FUNCTION_BLOCK "LKinCtrl_MC_ExecuteKinMotionCmd"   // FB35003, SCL
TITLE = LKinCtrl_ExecuteKinMotinCmd
{ S7_Optimized_Access := 'TRUE' }
AUTHOR : tech.team.motioncontrol@siemens.com
FAMILY : LKinCtrl
VERSION : 3.0
// FB executing single motion commands for TO_Kinematics. 
// - handling internal motion command instances
// - managing MotionQueue to be full, but not overloaded
// - providing status information on execution status
   VAR_INPUT
      execute : Bool;   // rising edge starts action once
      interrupt : Bool;   // trigger GroupInterrupt [interrupt input of FB_MovePath]
      continueMotion : Bool;   // trigger GroupContinue [no use in FB_MovePath] (used for FB_ExecutePathMotion stand alone)
      stop : Bool;   // trigger GroupStop [stop input of FB_MovePath]
      stopMode : DInt;   // MC_GroupStop dynamics; 0: stop with dynamics of active motion job; 1: stop with maximum kinematics dynamics (dynamics adaption still effective)
      reset : Bool;   // reset FB / acknowledge errors [reset input of FB_MovePath]
      writtenActiveCmdNo : DInt;   // last active cmdNo handled by FB MovePath
      conveyorConfiguration : Array[1.."LKINCTRL_NO_OF_CONVEYOR"] of "LKinCtrl_typeConveyorConfiguration";   // conveyor configuration / Conveyor configuration
   END_VAR
   VAR_OUTPUT
      done : Bool;   // TRUE: Commanded functionality has been completed successfully
      busy : Bool;   // TRUE: FB is not finished and new output values can be expected
      active : Bool;   // FB in control of axesGroup / kinematic in motion
      error : Bool;   // TRUE: An error occurred during the execution of the FB
      commandAborted : Bool;   // TRUE: Commanded functionality has been aborted by another command
      activePathDataName : String["LKINCTRL_LENGTH_OF_PATHDATA_NAME"];   // name of actual PathData
      activePathDataIdentifier : USInt;   // identifier number of actual PathData
      activeCmdNo : DInt;   // number of actual PathData set number
      cmdExecuted : Bool;   // actual pathData cmd executed to MotionQueue
      remainingDistanceActCmd : LReal;   // remainingDistance of active motionCommand
      waitTimeActive : Bool;   // TRUE: waitTime active in FB
      diagnostics : "LKinCtrl_typeExecuteKinMotionCmdDiagnostics";   // Diagnostics information of FB
   END_VAR
   VAR_IN_OUT
      pathDataElementPreBuf : "LKinCtrl_typePathDataElement_PreBuf";   // reference to the PathData element to be executed by FB_ExecuteKinMotionCmd
      to_Kinematics : TO_Kinematics;   // reference to the axesGroup
   END_VAR
   VAR
      statExecuteOld : Bool;   // old value of 'execute' input for edge detection
      statStopOld : Bool;   // old value of 'stop' input for edge detection
      statInterruptOld : Bool;   // old value of 'interrupt' input for edge detection
      statContinueMotionOld : Bool;   // old value of 'continueMotion' input for edge detection
      statResetOld : Bool;   // old value of 'reset' input for edge detection
      statDone : Bool;   // static value for output 'done'
      statBusy : Bool;   // static value for output 'busy'
      statCommandAborted : Bool;   // static value for output 'commandAborted'
      statActive : Bool;   // static value for output 'active'
      statActiveCmdNo : DInt;   // static value for output 'activeCmdNo'
      statWaitTimeActive : Bool;   // static value for output 'waitTimeActive'
      statWaitTime : Time;   // static time storage for time to wait for during wait time
      statError : Bool;   // static value for output 'error'
      statStatus : Word := 16#7000;   // static value for output 'status'
      statSubfunctionStatus : Word;   // Status or return value of called FBs, FCs and system blocks
      statFBState : Int := 0;   // State in the state machine of the FB
      statStateMachine : Int;   // static state machine status
      statDebugState : Bool;   // debug state machine by single steps
      statDebugFaultyValue : Int;   // debugging static for development only
      statDebugMessage : String;   // debugging string for development only
      statCmdExecuted : Bool;   // static value for output 'cmdExecuted'
      statExecWaitTime : Bool;   // execute flag for triggering wait time
      statExecFlagOnly : Bool;   // 'execute' flag for flagOnly dummy command
      statExecGroupInterrupt : Bool;   // execute flag for triggering MC_GroupInterrupt
      statExecGroupContinue : Bool;   // execute flag for triggering MC_GroupContinue
      statExecGroupStop : Bool;   // execute flag for triggering MC_GroupStop
      statExternalStopDetected : Bool;   // static storing informatioin on external stop being triggered
      statExecuteFlagOnlyCmd : Bool;   // static 'trigger' for execution of flag only cmd
      statStartCmdIsFlagOnly : Bool;   // static to store information that first command in PathData is flag only command
      statCmdIsMotionCmd : Bool;   // static containing cmd category; TRUE: motion cmd; FALSE: non-motion cmd
      statFBCounterLin : Int := 1;   // counter for organization of used linear motion FB instances
      statFBCounterCirc : Int := 1;   // counter for organization of used circular motion FB instances
      statFBCounterMoveDir : Int := 1;   // counter for organization of used move direct motion FB instances
      statFBCounterTrackConv : Int := 1;   // counter for organization of used conveyor tracking FB instances / counter for organization of used move direct motion FB instances
      statCoordSystemOld : DInt := 0;   // static storing old coordSystem information
      statLinkConstellation : DInt;   // static storing the link constellation
      statActualTrackedOCS : SInt;   // actually tracked OCS from kinematics
      statOCSInSync : SInt;   // OCS which is or will be syncrhonized to
      statBlendingRadius : LReal;   // calculated blending radius for SPTP commands
      statOCSInTracking : Array[1..3] of Bool;   // signalizes if a OCS is or will be used for tracking
      statLastPos : Array[1..4] of LReal;   // static for last TO_Kinematic position (for conversion relative to absolute motion)
      statAbsolutePosition : Array[1..4] of LReal;   // flag for AbsoultePosition of linear command to be changed internally (for conversion relative to absolute motion)
      statAuxPoint : Array[1..3] of LReal;   // flag for AuxPoint of circular command to be changed internally (for conversion relative to absolute motion)
      statEndPoint : Array[1..4] of LReal;   // flag for last EndPoint of circular command to be changed internally (for conversion relative to absolute motion)
      statExecLinCmds : Array[1..#LKINCTRL_MAX_NUMBER_OF_CMDS_LIN] of Bool;   // array of execute flags for triggering linear motion command FBs
      statExecCircCmds : Array[1..#LKINCTRL_MAX_NUMBER_OF_CMDS_CIRC] of Bool;   // array of execute flags for triggering circular motion command FBs
      statExecMoveDirectCmds : Array[1..#LKINCTRL_MAX_NUMBER_OF_CMDS_MOVEDIRECT] of Bool;   // array of execute flags for triggering move direct motion command FBs
      statExecTrackConv : Array[1..#LKINCTRL_MAX_NUMBER_OF_CMDS_TRACKCONV] of Bool;   // array of execute flags for triggering conveyor tracking command FBs / array of execute flags for triggering linear motion command FBs
      statConveyorBeltAxis : Array[1..#LKINCTRL_MAX_NUMBER_OF_CMDS_TRACKCONV] of DB_ANY;   // array of conveyor belt axes to be used at the instances
      statOCSFrames : Array[1..3] of "LKinCtrl_typeFrame";   // array of OCS frames
      statEmptyDiagnostics : "LKinCtrl_typeExecuteKinMotionCmdDiagnostics";   // empty diagnostics information (for initialization purposes only)
      statStoreExecuteBuffer : Struct   // struct for assignment of motion command FB instances PathData set specific data (setNo, PathDataNo)
         writeBufferElement : Int := 1;   // flag for set to be executed to MotionQueue in ExecuteBuffer struct
         activeBufferElement : Int := 1;   // flag for active set in ExecuteBuffer struct
         lastBufferElement : Int := 20;
         bufferElement : Array[1..#LKINCTRL_EXECUTEBUFFER_LENGTH] of Struct   // assignment of motion command FB instances PathData set specific data (setNo, PathDataNo)
            pathDataName : String["LKINCTRL_LENGTH_OF_PATHDATA_NAME"];
            pathDataIdentifier : USInt;
            setNumber : DInt;
            MotionFBNo : Int;
         END_STRUCT;
      END_STRUCT;
      statDebugExecCmdLogger : Struct   // command logger structure to store all executed commands (to MotionQueue), never deleted
         loggerElement : Array[1..#CONST_LENGTH_DATALOGGER] of Struct   // logger array storing executed commands and specific debug data
            executedCmd : "LKinCtrl_typeCmdLoggerElement";   // command
            executeBufferElement : Int;   // statStoreExecuteBuffer element number
            assignedMotionFB : Int;   // MC instance assigned
            timeStamp : Date_And_Time;   // time stamp of execution time of logged command
         END_STRUCT;
         writeCmdLoggerElement : Int := 1;   // pointer for writing logger element; incremented after writing ==> value -1 is last written element
         activeCmdLoggerElement : Int := 1;   // pointing on active cmd in command logger; showing active element during execution ==> after SUCCESSFUL completion of path incrementation ==> value -1 is last active element
      END_STRUCT;
      instMC_MoveLinAbs : Array[1..#LKINCTRL_MAX_NUMBER_OF_CMDS_LIN] of MC_MOVELINEARABSOLUTE;   // multi instance array MC_MoveLinearAbsoulte
      instMC_MoveCircAbs : Array[1..#LKINCTRL_MAX_NUMBER_OF_CMDS_CIRC] of MC_MOVECIRCULARABSOLUTE;   // multi instance array MC_MoveCircularAbsoulte
      instMC_MoveDirectAbs : Array[1..#LKINCTRL_MAX_NUMBER_OF_CMDS_MOVEDIRECT] of MC_MOVEDIRECTABSOLUTE;   // multi instance array MC_MoveDirectAbsoulte
      instMC_GROUPINTERRUPT : MC_GROUPINTERRUPT;   // multi instance MC_GroupInterrupt
      instMC_GROUPSTOP : MC_GROUPSTOP;   // multi instance FB MC_GroupStop
      instMC_GROUPCONTINUE : MC_GROUPCONTINUE;   // multi instance FB MC_GroupContinue
      instMC_KinematicsTransformation : MC_KINEMATICSTRANSFORMATION;   // multi instance FB MC_KinematicsTransformation
      instMC_InverseKinematicsTransformation : MC_INVERSEKINEMATICSTRANSFORMATION;   // multi instance FB MC_InverseKinematicsTransformation
      instMC_TrackConveyor : Array[1..3] of MC_TRACKCONVEYORBELT;   // multi instance FB MC_TrackConveyorBelt
      instIEC_Timer_waitTime : TON_TIME;   // multi instance TIMER_ON for wait times
   END_VAR
   VAR_TEMP
      tempExecute : Bool;   // Temporary value for input 'execute'
      tempStop : Bool;   // Temporary value for input 'stop'
      tempStopMode : DInt;   // Temporary value for input 'stopMode'
      tempInterrupt : Bool;   // Temporary value for input 'interrupt'
      tempContinueMotion : Bool;   // Temporary value for input 'continueMotion'
      tempReset : Bool;   // Temporary value for input 'reset'
      tempPosElemCtr : Int;   // Temporary counter variable
      tempCtr : Int;   // Temporary counter variable
      tempFBInstCtr : Int;   // Temporary counter variable
      tempMCActive : Bool;   // Temporary value to signal active MC instance
      tempMCBusy : Bool;   // Temporary value to signal busy MC instance
      tempRetVal : Int;   // Temporary return value
      tempRetValWord : Word;   // Temporary return value
      tempCmdType : Int;   // Temporary variable for type of command
      tempActiveInstance : Int;   // Temporary variable for active MC instance
      tempCmdDone : Bool;   // Temporary bit to signal done of MC instance
      tempCalc : Array[1..4] of LReal;   // Temporary calculation variable
      tempBlending : Array[1..4] of LReal;   // Temporary calculation variable
   END_VAR
   VAR CONSTANT
      NO_PROCESSING : Int := 0;   // FB_ExecutePathMotion state machine constant
      RESETTING : Int := 5;   // FB_ExecutePathMotion state machine constant
      RECEIVE_CMD : Int := 10;   // FB_ExecutePathMotion state machine constant
      CMD_CALC_SELECT : Int := 30;   // FB_ExecutePathMotion state machine constant
      EXEC_LIN : Int := 40;   // FB_ExecutePathMotion state machine constant
      EXEC_CIRC : Int := 41;   // FB_ExecutePathMotion state machine constant
      EXEC_MOVE_DIRECT : Int := 42;   // FB_ExecutePathMotion state machine constant
      EXEC_TRACK_CONV : Int := 43;   // FB_ExecutePathMotion state machine constant
      EXEC_SET_WS_ZONE : Int := 49;   // FB_ExecutePathMotion state machine constant
      EXEC_FLAG_ONLY : Int := 55;   // FB_ExecutePathMotion state machine constant
      EXEC_WAIT_TIME : Int := 57;   // FB_ExecutePathMotion state machine constant
      WAITING_TIME : Int := 58;   // FB_ExecutePathMotion state machine constant
      QUEUE_BUSY : Int := 60;   // FB_ExecutePathMotion state machine constant
      INTERRUPTING : Int := 70;   // FB_ExecutePathMotion state machine constant
      INTERRUPTED : Int := 75;   // FB_ExecutePathMotion state machine constant
      CONTINUEING : Int := 77;   // FB_ExecutePathMotion state machine constant
      CONTINUED : Int := 78;   // FB_ExecutePathMotion state machine constant
      STOPPING : Int := 80;   // FB_ExecutePathMotion state machine constant
      STOPPED_STATE : Int := 85;   // FB_ExecutePathMotion state machine constant
      DESYNC_CONVEYOR : Int := 86;   // FB_ExecutePathMotion state machine constant
      ERROR_STATE : Int := 90;   // FB_ExecutePathMotion state machine constant
      LKINCTRL_MAX_NUMBER_OF_CMDS_LIN : Int := 12;   // max number of MC_MoveLinearAbsolute FB instances
      LKINCTRL_MAX_NUMBER_OF_CMDS_CIRC : Int := 12;   // max number of MC_MoveCircularAbsolute FB instances
      LKINCTRL_MAX_NUMBER_OF_CMDS_MOVEDIRECT : Int := 12;   // max number of MC_MoveDirectAbsolute FB instances
      LKINCTRL_MAX_NUMBER_OF_CMDS_TRACKCONV : Int := 3;   // max number of MC_TrackConveyorBelt FB instances
      LKINCTRL_EXECUTEBUFFER_LENGTH : Int := 12;   // length of internal buffer (needs to be set to same value as LKINCTRL_MAX_NUMBER_OF_CMDS_LIN)
      STATUS_NO_ERROR : Word := 16#0000;   // status no error
      STATUS_NO_CALL : Word := 16#7000;   // No job being currently processed
      STATUS_FIRST_CALL : Word := 16#7001;   // First call after incoming new job (rising edge 'execute')
      STATUS_SUBSEQUENT_CALL : Word := 16#7002;   // Subsequent call during active processing without further details
      STATUS_CMD_EXECUTED : Word := 16#7010;   // status command executed to MotionQueue
      STATUS_PATHMOTION_RUNNING : Word := 16#7100;   // status path motion running
      STATUS_PATHMOTION_INTERRUPTING : Word := 16#7101;   // status path motion interrupting
      STATUS_PATHMOTION_INTERRUPTED : Word := 16#7102;   // status path motion interrupted
      STATUS_PATHMOTION_STOPPING : Word := 16#7103;   // status path motion stopping
      STATUS_COMMAND_ABORTED : Word := 16#7104;   // commanded functionality has been aborted by another command
      STATUS_PATHMOTION_CONTINUEING : Word := 16#7105;   // status path motion continueing
      STATUS_FB_RESETTING : Word := 16#7106;   // status FB reset
      STATUS_WAIT_TIME_ACTIVE : Word := 16#7107;   // status wait time active
      STATUS_WAIT_TIME_FINISHED : Word := 16#7108;   // status wait time finished
      STATUS_PATHMOTION_EXT_STOPPING : Word := 16#7109;   // status external stop active
      STATUS_PATHMOTION_BUFFER_BUSY : Word := 16#7111;   // status motionQueue full / buffer busy
      STATUS_PATHMOTION_FINISHED : Word := 16#7110;   // status path motion finished / end of path position reached
      STATUS_DESYNC_CONVEYOR : Word := 16#7112;   // status desync from conveyor with motion command
      ERR_UNDEFINED_STATE : Word := 16#8600;   // error due to an undefined state in state machine
      ERR_GROUPINTERRUPT_FAILED : Word := 16#8242;   // error MC_GroupInterrupt failed
      ERR_GROUPCONTINUE_FAILED : Word := 16#8243;   // error MC_GroupContinue failed
      ERR_GROUPSTOP_FAILED : Word := 16#8244;   // error MC_GroupStop failed
      ERR_TO_KINEMATIC_ERROR : Word := 16#8245;   // error in TO_Kinematic
      ERR_LINEAR_CMD : Word := 16#8246;   // error MC_MoveLinear failed
      ERR_CIRCULAR_CMD : Word := 16#8247;   // error MC_MoveCircular failed
      ERR_CMD_PARAMETER : Word := 16#8248;   // error command parametrization
      ERR_CALC_CIRC_CMD : Word := 16#8249;   // error circular command conversion: arc calculation
      ERR_MOVEDIRECT_CMD : Word := 16#8250;   // error MC_MoveDirect failed
      ERR_TRACKCONVEYOR_CMD : Word := 16#8251;   // error MC_TrackConveyorBelt failed
      ERR_DESYNC_RELATIVE : Word := 16#8252;   // error due to relative command used for desync conveyor
      ERR_CONVEYOR_CONFIGURATION : Word := 16#8253;   // error due to invalid conveyor configuration
      CONST_LENGTH_DATALOGGER : Int := 15;   // length of internal data logger
      SPTP_REMAINING_DIST : Bool := FALSE;   // TRUE: Caclulate own RemainingDistance for SPTP / FALSE: Use ExecutionTimeStatus
      SPTP_APPROX_BLENDING : Bool := FALSE;   // TRUE: When remDistance is calculated also approximate blending distance / FALSE: Set blending is not regarded on calculation
   END_VAR
   // statStoreExecuteBuffer.bufferElement[12].MotionFBNo := -1;
   // statStoreExecuteBuffer.bufferElement[11].MotionFBNo := -1;
   // statStoreExecuteBuffer.bufferElement[10].MotionFBNo := -1;
   // statStoreExecuteBuffer.bufferElement[9].MotionFBNo := -1;
   // statStoreExecuteBuffer.bufferElement[8].MotionFBNo := -1;
   // statStoreExecuteBuffer.bufferElement[7].MotionFBNo := -1;
   // statStoreExecuteBuffer.bufferElement[6].MotionFBNo := -1;
   // statStoreExecuteBuffer.bufferElement[5].MotionFBNo := -1;
   // statStoreExecuteBuffer.bufferElement[4].MotionFBNo := -1;
   // statStoreExecuteBuffer.bufferElement[3].MotionFBNo := -1;
   // statStoreExecuteBuffer.bufferElement[2].MotionFBNo := -1;
   // statStoreExecuteBuffer.bufferElement[1].MotionFBNo := -1;
   // statDebugExecCmdLogger.loggerElement[10].assignedMotionFB := -1;
   // statDebugExecCmdLogger.loggerElement[10].executeBufferElement := -1;
   // statDebugExecCmdLogger.loggerElement[9].assignedMotionFB := -1;
   // statDebugExecCmdLogger.loggerElement[9].executeBufferElement := -1;
   // statDebugExecCmdLogger.loggerElement[8].assignedMotionFB := -1;
   // statDebugExecCmdLogger.loggerElement[8].executeBufferElement := -1;
   // statDebugExecCmdLogger.loggerElement[7].assignedMotionFB := -1;
   // statDebugExecCmdLogger.loggerElement[7].executeBufferElement := -1;
   // statDebugExecCmdLogger.loggerElement[6].assignedMotionFB := -1;
   // statDebugExecCmdLogger.loggerElement[6].executeBufferElement := -1;
   // statDebugExecCmdLogger.loggerElement[5].assignedMotionFB := -1;
   // statDebugExecCmdLogger.loggerElement[5].executeBufferElement := -1;
   // statDebugExecCmdLogger.loggerElement[4].assignedMotionFB := -1;
   // statDebugExecCmdLogger.loggerElement[4].executeBufferElement := -1;
   // statDebugExecCmdLogger.loggerElement[3].assignedMotionFB := -1;
   // statDebugExecCmdLogger.loggerElement[3].executeBufferElement := -1;
   // statDebugExecCmdLogger.loggerElement[2].assignedMotionFB := -1;
   // statDebugExecCmdLogger.loggerElement[2].executeBufferElement := -1;
   // statDebugExecCmdLogger.loggerElement[1].assignedMotionFB := -1;
   // statDebugExecCmdLogger.loggerElement[1].executeBufferElement := -1;
BEGIN
   //==========================================================================================
   // SIEMENS AG
   // (c)Copyright 2020 All Rights Reserved
   //------------------------------------------------------------------------------------------
   // Library: LKinCtrl
   // Tested with: S7-1517T-3 PN/DP
   // Engineering: TIA Portal V16
   // Restrictions: ---
   // Requirements: S7-1500T FW 2.8
   // Functionality: LKinCtrl_MC_ExecuteKinMotionCmd
   // The FB is executing the motion commands requested and received from the
   // PathDataPreBuffered structure. The TO_Kinematics motion queue is kept busy and command
   // buffering is managed not to exceed motion queues limits.
   // 
   // Support: tech.team.motioncontrol@siemens.com
   // Note: Parameter comments are only available in language 'English (United States)'
   //------------------------------------------------------------------------------------------
   // Change log table:
   // Version    Date          Expert in charge    Changes applied
   // 01.00.00   06.02.2018    JR                  First release version V1.0
   // 02.00.00   18.04.2019    JR / FR             V2.0
   // 02.00.01   29.04.2019    JR                  fix for relative circle last pos calc
   // 02.00.02   03.05.2019    FR                  added ParameterValid bits
   // 02.01.00   28.05.2019    JR / FR             V2.1 for LKinLang
   // 02.02.00   28.01.2020    JR / FR             V2.2: Added valueFlags and flagOnlyCmd 
   // 02.02.01   07.02.2020    FR / DF             V2.2.1: Fix of active output in case of circular commands and fix of activeBufferElement when path motion is finished
   // 02.03.00   18.03.2020    FR                  Fix for interrupt / continue; Added static for "active" and "waitTimeActive" output
   // 02.03.01   14.04.2020    FR                  Bugfixes and partial rework
   // 02.03.02   16.07.2020    FR                  Bugfixes
   // 03.00.00   04.08.2020    FR                  Added MoveDirect and ConveyorTracking; Bugfixes and partial rework
   // 03.00.01   07.08.2020    FR                  Bugfix for WaitTime timing
   // 03.00.02   19.10.2020    FR                  Workaround for stop when command finishes; Workaround for MC_TrackConveyorBelt; Only update activeCmdNo if cmd is actually active
   // 03.00.03   15.12.2020    FR                  Reset static when ending with flag command; Bugfix for interrupt / continue; added RemainingDistance calculation for SPTP
   // 03.00.04   06.07.2021    FR                  Bugfix for interrupt / continue
   //===========================================================================================

   // Work with temporary values / create process images
   #tempExecute := #execute;
   #tempStop := #stop;
   #tempInterrupt := #interrupt;
   #tempContinueMotion := #continueMotion;
   #tempReset := #reset;
   #tempStopMode := #stopMode;

   REGION TRIGGERING
     //===========================================================================================
     // check for risind edge of stop input
     IF (#tempStop = TRUE) AND (#statStopOld = FALSE)
     THEN
       // FR 29.04.2020: Set FB busy when stopping! 
       #statBusy := TRUE;
       #statDone := FALSE;
       #statCommandAborted := FALSE;
       #statError := FALSE;

       // perform stop procedure
       #statStateMachine := #STOPPING;
       // set status accordingly
       #statStatus := #STATUS_PATHMOTION_STOPPING;
       //===========================================================================================
       // check for risind edge of interrupt input
     ELSIF (#tempInterrupt = TRUE) AND (#statInterruptOld = FALSE)
     THEN
       // perform interrupt procedure
       #statStateMachine := #INTERRUPTING;
       // set status according
       #statStatus := #STATUS_PATHMOTION_INTERRUPTING;
       //===========================================================================================
       // check for risind edge of continueMotion input
     ELSIF (#tempContinueMotion = TRUE) AND (#statContinueMotionOld = FALSE)
     THEN
       // perform continue procedure
       #statStateMachine := #CONTINUEING;
       // set status accordingly
       #statStatus := #STATUS_PATHMOTION_CONTINUEING;
       //===========================================================================================
       // check for risind edge of reset input
     ELSIF (#tempReset = TRUE) AND (#statResetOld = FALSE)
       // interlock reset during execution
       AND (#statBusy = FALSE)
     THEN
       // perform reset procedure
       #statStateMachine := #RESETTING;
       // set status accordingly
       #statStatus := #STATUS_FB_RESETTING;
       //===========================================================================================
       // check for risind edge of execute input
     ELSIF (#tempExecute = TRUE) AND (#statExecuteOld = FALSE)
       // interlock input signals at stop / interrupt / reset
       AND (#stop = FALSE) AND (#interrupt = FALSE) AND (#reset = FALSE)
       // interlock triggering during WAIT_TIME active or waiting to be active
       AND (#statStateMachine <> #EXEC_WAIT_TIME) AND (#statStateMachine <> #WAITING_TIME)
     THEN
       // First call; initialize FB
       #statDone := FALSE;
       #statBusy := TRUE;
       #statCommandAborted := FALSE;
       // #statError := FALSE;
       #statStatus := #STATUS_FIRST_CALL;

       // FR 25.06.2020: Commented to allow interrupt and filling of queue
       // //------------------------------------------------------------------------------------------
       // // check for TO Kinematics to be interrupted ==> continue path
       // IF #to_Kinematics.StatusWord.%X17
       //     AND #statStateMachine = #INTERRUPTED
       // THEN
       //     #statStateMachine := #CONTINUEING;
       //     #statStatus := #STATUS_PATHMOTION_CONTINUEING;
       //     //------------------------------------------------------------------------------------------
       //     // check for already pending error ==> do nothing in case of error
       // ELS
       IF #statError THEN
         #statStateMachine := #ERROR_STATE;
         //------------------------------------------------------------------------------------------
         // start processing
         // check for TO Kinematics not to be interrupted and no error pending
       ELSE
         // set state machine to starting state
         #statStateMachine := #RECEIVE_CMD;

         // check for active MC linear instance
         FOR #tempCtr := 1 TO #LKINCTRL_MAX_NUMBER_OF_CMDS_LIN DO
           IF #instMC_MoveLinAbs[#tempCtr].Execute THEN
             // set temp to interlock reset
             #tempMCActive := TRUE;
             EXIT;
           ELSE
             #tempMCActive := FALSE;
           END_IF;
         END_FOR;
         // check for no circular instance to be busy in case of no linear cmd busy
         IF #tempMCActive = FALSE THEN
           FOR #tempCtr := 1 TO #LKINCTRL_MAX_NUMBER_OF_CMDS_CIRC DO
             IF #instMC_MoveCircAbs[#tempCtr].Execute THEN
               // set temp to interlock reset
               #tempMCActive := TRUE;
               EXIT;
             ELSE
               #tempMCActive := FALSE;
             END_IF;
           END_FOR;
         END_IF;
         // check for no PTP instance to be busy in case of no linear cmd busy
         IF #tempMCActive = FALSE THEN
           FOR #tempCtr := 1 TO #LKINCTRL_MAX_NUMBER_OF_CMDS_MOVEDIRECT DO
             IF #instMC_MoveDirectAbs[#tempCtr].Execute THEN
               // set temp to interlock reset
               #tempMCActive := TRUE;
               EXIT;
             ELSE
               #tempMCActive := FALSE;
             END_IF;
           END_FOR;
         END_IF;

         // initialization of variables - in stillstand and with no command active only
         IF #to_Kinematics.StatusMotionQueue.NumberOfCommands = 0
           AND #to_Kinematics.StatusPath.Velocity = 0.0
           // AND #to_Kinematics.StatusWord.%X17 = FALSE    // double check for TO interrupted ==> could be removed ?!
           // AND #to_Kinematics.StatusWord.%X6 = TRUE   // no job active on TO Kinematics
           AND #to_Kinematics.StatusWord.%X8 = FALSE     // no linear command active on TO Kinematics
           AND #to_Kinematics.StatusWord.%X9 = FALSE     // no cicrular command active on TO Kinematics
           AND #to_Kinematics.StatusWord.%X11 = FALSE    // no moveDirect command active on TO Kinematics
           AND #instIEC_Timer_waitTime.ET = t#0ms        // no timer running
           AND #tempMCActive = FALSE                     // none of the MC instances busy, in case of asymmetric signal of instance.busy & TO_Kinematics.X6 (job done)
           AND #statExecuteFlagOnlyCmd = FALSE           // no flag only command 'active' (activeCmdNo visible for one cycle, no initialization in that cycle !)
         THEN
           // reset FB counters for MC command instances
           #statFBCounterLin := 1;
           #statFBCounterCirc := 1;
           #statFBCounterMoveDir := 1;
           //#statFBCounterTrackConv := 1; // 07.08.2020 FR: Use every instance of MC_TrackConveyor
           // Reset blending radius calculation
           #statBlendingRadius := -1;
           // reset all execute triggers of motion commands
           FOR #tempCtr := 1 TO #LKINCTRL_MAX_NUMBER_OF_CMDS_LIN DO
             #statExecLinCmds[#tempCtr] := FALSE;
             #statExecCircCmds[#tempCtr] := FALSE;
             #statExecMoveDirectCmds[#tempCtr] := FALSE;
           END_FOR;

           FOR #tempCtr := 1 TO #LKINCTRL_MAX_NUMBER_OF_CMDS_TRACKCONV DO
             #statExecTrackConv[#tempCtr] := FALSE;
           END_FOR;

           // Reset waitTimer execute
           #statExecWaitTime := FALSE;

           // Reset instances
           #instMC_InverseKinematicsTransformation(AxesGroup := #to_Kinematics,
                                                   Enable := FALSE);
           #instMC_KinematicsTransformation(AxesGroup := #to_Kinematics,
                                            Enable := FALSE);

           // reset store buffer variables for handling activeCmdNo assigment
           #statStoreExecuteBuffer.writeBufferElement := 0;//1;
           #statStoreExecuteBuffer.activeBufferElement := 1;
           // synchronize data logger active and write element
           #statDebugExecCmdLogger.activeCmdLoggerElement := #statDebugExecCmdLogger.writeCmdLoggerElement;
           FOR #tempCtr := 1 TO #LKINCTRL_EXECUTEBUFFER_LENGTH DO
             #statStoreExecuteBuffer.bufferElement[#tempCtr].pathDataName := '';
             #statStoreExecuteBuffer.bufferElement[#tempCtr].setNumber := 0;
             #statStoreExecuteBuffer.bufferElement[#tempCtr].MotionFBNo := -1;
           END_FOR;

           // Get initial position
           // WCS
           #statLastPos[1] := #to_Kinematics.Tcp.x;
           #statLastPos[2] := #to_Kinematics.Tcp.y;
           #statLastPos[3] := #to_Kinematics.Tcp.z;
           #statLastPos[4] := #to_Kinematics.Tcp.a;
           // reset old coordinate system information
           #statCoordSystemOld := "CS_WCS";

           // Get initial link constellation
           #statLinkConstellation := DWORD_TO_DINT(#to_Kinematics.StatusKinematics.LinkConstellation);

           // Added FR: 2020/01/27
           // Check if next cmdId is higher than active cmd --> Assume path is continued after wait flag/time
           IF #pathDataElementPreBuf.cmdID > #statActiveCmdNo THEN
             // Do not reset activeCmdNo --> 0 would appear on MovePath output
             ;
           ELSE
             // Reset activeCmdNo at beginning of new path data
             // added JR: 2019/11/27
             // reset output for activeCmd information
             #statActiveCmdNo := 0;
             #activePathDataName := '';
           END_IF;

           #remainingDistanceActCmd := 0.0;
           // reset flagOnly command storage bit
           #statExecuteFlagOnlyCmd := FALSE;
           // detect PathData starting with flagOnly command (not for readyForNextPath)
           IF #pathDataElementPreBuf.cmdType = "LKINCTRL_CMD_FLAG_ONLY" THEN
             // Statement section IF
             #statStartCmdIsFlagOnly := TRUE;
           ELSE
             #statStartCmdIsFlagOnly := FALSE;
           END_IF;

         END_IF;
         // initialization of variables - also while in motion
         #statCmdExecuted := FALSE;
         #statExecGroupStop := FALSE;
         #statExecGroupContinue := FALSE;
         #statExecGroupInterrupt := FALSE;
         #statExternalStopDetected := FALSE;
         #diagnostics := #statEmptyDiagnostics;
       END_IF;
       //------------------------------------------------------------------------------------------

       // initialization of variables
       #statCmdExecuted := FALSE;

     ELSIF (#statStatus = #STATUS_FIRST_CALL) THEN
       #statStatus := #STATUS_SUBSEQUENT_CALL;
     END_IF;

     // Edge detection input variables
     #statExecuteOld := #tempExecute;
     #statStopOld := #tempStop;
     #statInterruptOld := #tempInterrupt;
     #statContinueMotionOld := #tempContinueMotion;
     #statResetOld := #tempReset;

   END_REGION TRIGGERING

   IF (#statStatus = #STATUS_NO_CALL) THEN // Nothing to do -> End here to reduce "system load"
     // RETURN;
     ;
   END_IF;

   REGION STATE_MACHINE

     // no processing state ==> do nothing
     REGION NO_PROCESSING
       IF #statStateMachine = #NO_PROCESSING
         // AND #statDebugState = TRUE
       THEN
         // reset  variable for single step debugging of states
         #statDebugState := FALSE;
         // do nothing
         ;
       END_IF;
     END_REGION NO_PROCESSING

     // state reached when reset is executed
     REGION RESETTING
       IF #statStateMachine = #RESETTING
         // AND #statDebugState = TRUE
       THEN
         // reset  variable for single step debugging of states
         #statDebugState := FALSE;

         // reset state machine
         #statStateMachine := #NO_PROCESSING;

         // reset FB counters for MC command instances
         #statFBCounterLin := 1;
         #statFBCounterCirc := 1;
         #statFBCounterMoveDir := 1;
         #statFBCounterTrackConv := 1;
         // Reset blending radius calculation
         #statBlendingRadius := -1;
         // reset all execute triggers of motion commands
         FOR #tempCtr := 1 TO #LKINCTRL_MAX_NUMBER_OF_CMDS_LIN DO
           #statExecLinCmds[#tempCtr] := FALSE;
           #statExecCircCmds[#tempCtr] := FALSE;
           #statExecMoveDirectCmds[#tempCtr] := FALSE;
         END_FOR;

         FOR #tempCtr := 1 TO #LKINCTRL_MAX_NUMBER_OF_CMDS_TRACKCONV DO
           #statExecTrackConv[#tempCtr] := FALSE;
         END_FOR;

         // Reset instances
         #instMC_InverseKinematicsTransformation(AxesGroup := #to_Kinematics,
                                                 Enable := FALSE);
         #instMC_KinematicsTransformation(AxesGroup := #to_Kinematics,
                                          Enable := FALSE);

         // reset store buffer variables for handling activeCmdNo assigment
         #statStoreExecuteBuffer.writeBufferElement := 0;//1;
         #statStoreExecuteBuffer.activeBufferElement := 1;
         FOR #tempCtr := 1 TO #LKINCTRL_EXECUTEBUFFER_LENGTH DO
           #statStoreExecuteBuffer.bufferElement[#tempCtr].pathDataName := '';
           #statStoreExecuteBuffer.bufferElement[#tempCtr].setNumber := 0;
           #statStoreExecuteBuffer.bufferElement[#tempCtr].MotionFBNo := -1;
         END_FOR;
         // reset static variables for output signals
         #statCmdExecuted := FALSE;
         #statExecGroupStop := FALSE;
         #statExecGroupContinue := FALSE;
         #statExecGroupInterrupt := FALSE;
         #statExecWaitTime := FALSE;
         #statExternalStopDetected := FALSE;
         #statCoordSystemOld := "CS_WCS";
         #diagnostics := #statEmptyDiagnostics;
         // reset output for activeCmd information
         #statActiveCmdNo := 0;
         #activePathDataName := '';
         #remainingDistanceActCmd := 0.0;
         // set status
         #statStatus := #STATUS_NO_CALL;
       END_IF;
     END_REGION RESETTING



     // reception of new commands from CmdHandler
     REGION RECEIVE_CMD
       IF #statStateMachine = #RECEIVE_CMD
         // AND #statDebugState = TRUE
       THEN
         // reset  variable for single step debugging of states
         #statDebugState := FALSE;

         // check for MotionQueue not to be full
         IF #to_Kinematics.StatusMotionQueue.NumberOfCommands < #to_Kinematics.MotionQueue.MaxNumberOfCommands
           AND (#statStoreExecuteBuffer.activeBufferElement <> #statStoreExecuteBuffer.writeBufferElement) // FR 09.06.2020: Do not overwrite active buffer element!
         THEN
           // Init writeBuffer to 1 if 0; only is 0 after reset or first cycle
           IF #statStoreExecuteBuffer.writeBufferElement = 0 THEN
             #statStoreExecuteBuffer.writeBufferElement := 1;
           END_IF;

           // check command parameters to be correct
           #statSubfunctionStatus := "LKinCtrl_CheckPathDataCmd"(cmdIsMotionCmd => #statCmdIsMotionCmd, pathDataCmd := #pathDataElementPreBuf);

           // Check if conveyor parameter if cmd is MC_TrackConveyorBelt
           IF #pathDataElementPreBuf.cmdType = "LKINCTRL_MC_TRACKCONVEYORBELT" THEN
             // Check axis DB number
             IF #conveyorConfiguration[#pathDataElementPreBuf.cmdParameters.conveyorParameters.conveyorParaNo].conveyorBeltAxis = 0 THEN
               // No axis connected --> Error
               #statStatus := #ERR_CONVEYOR_CONFIGURATION;

               // Check initial object position --> only x allowed
             ELSIF #conveyorConfiguration[#pathDataElementPreBuf.cmdParameters.conveyorParameters.conveyorParaNo].initialObjectPosition.y <> 0.0
               OR #conveyorConfiguration[#pathDataElementPreBuf.cmdParameters.conveyorParameters.conveyorParaNo].initialObjectPosition.z <> 0.0
               OR #conveyorConfiguration[#pathDataElementPreBuf.cmdParameters.conveyorParameters.conveyorParaNo].initialObjectPosition.a <> 0.0
               OR #conveyorConfiguration[#pathDataElementPreBuf.cmdParameters.conveyorParameters.conveyorParaNo].initialObjectPosition.b <> 0.0
               OR #conveyorConfiguration[#pathDataElementPreBuf.cmdParameters.conveyorParameters.conveyorParaNo].initialObjectPosition.c <> 0.0
             THEN
               // Initial object position not allowed --> Error
               #statStatus := #ERR_CONVEYOR_CONFIGURATION;
             END_IF;
           END_IF;

           // Check if desync from conveyor with relative command
           IF #pathDataElementPreBuf.cmdType = "LKINCTRL_MC_MOVELINEARREL"
             AND #statOCSInSync <> 0 // Check for conveyorTracking to be planned
             AND #pathDataElementPreBuf.cmdCoordinates.coordSystem <> #statOCSInSync
           THEN
             // Deysnc with relative command not allowed --> Error
             #statStatus := #ERR_DESYNC_RELATIVE;
           END_IF;

           IF #statSubfunctionStatus = #STATUS_NO_ERROR AND #statStatus.%X15 = FALSE THEN
             // new command not executed yet
             #statCmdExecuted := FALSE;
             // go to next state - command calculation and selection
             #statStateMachine := #CMD_CALC_SELECT;
           ELSIF #statSubfunctionStatus <> #STATUS_NO_ERROR THEN
             // new command not executed yet
             #statCmdExecuted := FALSE;
             // set status accordingly
             #statStatus := #ERR_CMD_PARAMETER;
             // set error information
             #diagnostics.faultSetNumber := #pathDataElementPreBuf.cmdID;
             #diagnostics.faultPathDataName := #pathDataElementPreBuf.pathDataName;
             // statSubFunctionStatus contains specific parameter error information (will be written at the bottom)
             // set state machine
             #statStateMachine := #ERROR_STATE;
           ELSIF #statStatus.%X15 THEN
             // new command not executed yet
             #statCmdExecuted := FALSE;
             // set error information
             #diagnostics.faultSetNumber := #pathDataElementPreBuf.cmdID;
             #diagnostics.faultPathDataName := #pathDataElementPreBuf.pathDataName;
             // statSubFunctionStatus contains specific parameter error information (will be written at the bottom)
             // set state machine
             #statStateMachine := #ERROR_STATE;
           END_IF;

         ELSE
           // continue in other state if MotionQueue is full
           #statStateMachine := #QUEUE_BUSY;
         END_IF;
       END_IF;
     END_REGION RECEIVE_CMD


     // calculation of command coordinates (conversion relative to absoulte) & command selection (linear or circular)
     REGION CMD_CALC_SELECT
       IF #statStateMachine = #CMD_CALC_SELECT
         // AND #statDebugState = TRUE
       THEN
         // reset  variable for single step debugging of states
         #statDebugState := FALSE;

         //------------------------------------------------------------------------------------------
         // Convert coordinates/command to absolute and check parameterValid bits
         //------------------------------------------------------------------------------------------
         IF #statCmdIsMotionCmd THEN // check for command type to be MC command (not WAIT_TIME or FlagOnly)
           //------------------------------------------------------------------------------------------
           // Transform statLastPos into correct CS
           //------------------------------------------------------------------------------------------
           // TODO: Integrate InverseKinTrans into FC LKinCtrl_FrameTrans ?
           IF #pathDataElementPreBuf.cmdCoordinates.coordSystem = "CS_MCS"
             AND #statCoordSystemOld <> "CS_MCS"
           THEN
             // Transform lastPos to MCS 
             #instMC_InverseKinematicsTransformation(AxesGroup := #to_Kinematics,
                                                     Enable := TRUE,
                                                     Position := #statLastPos,
                                                     CoordSystem := #statCoordSystemOld,
                                                     LinkConstellation := #statLinkConstellation,
                                                     ErrorId => #statSubfunctionStatus,
                                                     AxesPosition => #statLastPos);

           ELSIF #pathDataElementPreBuf.cmdCoordinates.coordSystem <> "CS_MCS"
             AND #statCoordSystemOld = "CS_MCS"
           THEN
             // Transform lastPos to target CS
             #instMC_KinematicsTransformation(AxesGroup := #to_Kinematics,
                                              Enable := TRUE,
                                              AxesPosition := #statLastPos,
                                              CoordSystem := #pathDataElementPreBuf.cmdCoordinates.coordSystem,
                                              ErrorId => #statSubfunctionStatus,
                                              Position => #statLastPos,
                                              LinkConstellation => #statLinkConstellation);

           ELSE
             // FR 29.04.2020: Update OCS frames every time in case they were changed
             FOR #tempCtr := 1 TO 3 DO
               #statOCSFrames[#tempCtr].x := #to_Kinematics.StatusOcsFrame[#tempCtr].x;
               #statOCSFrames[#tempCtr].y := #to_Kinematics.StatusOcsFrame[#tempCtr].y;
               #statOCSFrames[#tempCtr].z := #to_Kinematics.StatusOcsFrame[#tempCtr].z;
               #statOCSFrames[#tempCtr].a := #to_Kinematics.StatusOcsFrame[#tempCtr].a;
               #statOCSFrames[#tempCtr].b := #to_Kinematics.StatusOcsFrame[#tempCtr].b;
               #statOCSFrames[#tempCtr].c := #to_Kinematics.StatusOcsFrame[#tempCtr].c;
             END_FOR;

             // FR 26.03.2020: Updated FrameTrans 
             // Transform LastPos to correct CS
             "LKinCtrl_FrameTrans"(coordSystem := #pathDataElementPreBuf.cmdCoordinates.coordSystem, // Actual/Target CS
                                   coordSystemOld := #statCoordSystemOld, // Last CS
                                   OCSFrames := #statOCSFrames, // OCS frames
                                   position := #statLastPos); // Position to be transformed
           END_IF;

           // Check if KinTrans FBs returned no error
           IF #statSubfunctionStatus = #STATUS_NO_ERROR THEN
             // Update old CS
             #statCoordSystemOld := #pathDataElementPreBuf.cmdCoordinates.coordSystem;

             // Update tracked OCS 
             IF #statCoordSystemOld >= "CS_OCS1" AND #statCoordSystemOld <= "CS_OCS3" THEN
               IF #statOCSInTracking[#statCoordSystemOld] THEN
                 #statOCSInSync := DINT_TO_SINT(#statCoordSystemOld);
               END_IF;
             ELSIF #statCoordSystemOld = "CS_WCS" THEN
               #statOCSInSync := 0;
             END_IF;

             //------------------------------------------------------------------------------------------
             // Update linkConstellation
             //------------------------------------------------------------------------------------------
             // LinkConstellation can only be set at sPTP command in WCS/OCS
             IF #pathDataElementPreBuf.cmdCoordinates.coordSystem <> "CS_MCS"
               AND #pathDataElementPreBuf.cmdParameters.moveDirectParameters.linkConstellation <> 16#FFFF_FFFF
               AND (#pathDataElementPreBuf.cmdType = "LKINCTRL_MC_MOVEDIRECTABS"
               OR #pathDataElementPreBuf.cmdType = "LKINCTRL_MC_MOVEDIRECTREL")
             THEN
               // LinkConstellation is changed
               #statLinkConstellation := DWORD_TO_DINT(#pathDataElementPreBuf.cmdParameters.moveDirectParameters.linkConstellation);
             END_IF;

             //------------------------------------------------------------------------------------------
             // Update PositionMode
             //------------------------------------------------------------------------------------------
             // PositionMode is only valid for absolute SPTP command in WCS/OCS
             IF #pathDataElementPreBuf.cmdCoordinates.coordSystem <> "CS_MCS"
               AND #pathDataElementPreBuf.cmdParameters.moveDirectParameters.positionMode = 2 // Relative A coordinate
               AND #pathDataElementPreBuf.cmdType = "LKINCTRL_MC_MOVEDIRECTABS"
             THEN
               // Calc correct orientation position
               #statAbsolutePosition[4] := #statLastPos[4] + #pathDataElementPreBuf.cmdCoordinates.absolutePosition[4];
             END_IF;

             // Always set positionMode to 1 for absolute A Coordinate
             #pathDataElementPreBuf.cmdParameters.moveDirectParameters.positionMode := 1;

             //------------------------------------------------------------------------------------------
             // ParameterValid bit check
             //------------------------------------------------------------------------------------------
             IF #pathDataElementPreBuf.cmdType = "LKINCTRL_MC_MOVELINEARABS"
               OR #pathDataElementPreBuf.cmdType = "LKINCTRL_MC_MOVECIRCULARABS"
               OR #pathDataElementPreBuf.cmdType = "LKINCTRL_MC_MOVEDIRECTABS"
             THEN
               FOR #tempPosElemCtr := 1 TO "LKINCTRL_NO_OF_VALID_BITS" DO
                 // Check valid bits and copy last pos (X,Y,Z,A) where missing
                 IF #pathDataElementPreBuf.parameterValid[#tempPosElemCtr] = FALSE THEN
                   #pathDataElementPreBuf.cmdCoordinates.absolutePosition[#tempPosElemCtr] := #statLastPos[#tempPosElemCtr];
                 ELSE
                   ; // Keep programmed position from #pathDataElementPreBuf.cmdCoordinates.absolutePosition
                 END_IF;
               END_FOR;
             ELSIF #pathDataElementPreBuf.cmdType = "LKINCTRL_MC_MOVELINEARREL"
               OR #pathDataElementPreBuf.cmdType = "LKINCTRL_MC_MOVECIRCULARREL"
               OR #pathDataElementPreBuf.cmdType = "LKINCTRL_MC_MOVEDIRECTREL"
             THEN
               FOR #tempPosElemCtr := 1 TO "LKINCTRL_NO_OF_VALID_BITS" DO
                 // Check valid bits and set absolute pos to 0.0 (X,Y,Z,A)
                 IF #pathDataElementPreBuf.parameterValid[#tempPosElemCtr] = FALSE THEN
                   #pathDataElementPreBuf.cmdCoordinates.absolutePosition[#tempPosElemCtr] := 0.0;
                 ELSE
                   ; // Keep programmed position from #pathDataElementPreBuf.cmdCoordinates.absolutePosition
                 END_IF;
               END_FOR;
             ELSE
               ; // Nothing to do for this cmdType
             END_IF;

           ELSE
             // set error information
             #diagnostics.faultSetNumber := #pathDataElementPreBuf.cmdID;
             #diagnostics.faultPathDataName := #pathDataElementPreBuf.pathDataName;
             // statSubFunctionStatus contains error information (will be written at the bottom)
             // set state machine
             #statStateMachine := #ERROR_STATE;
           END_IF;